// TIA Portal project "PalletizerLine" (V17) (continued)
VERSION : 1.0
// Support: tech.team.motioncontrol@siemens.com
// Fax: +49 (0) 9131/98-1297
   VAR
      Summation : "CPG_typeEventSummation";   // Unit Mode - PackML Event Summation
   END_VAR
BEGIN
   Summation.wrk_EventArraySize := 30;
END_DATA_BLOCK

DATA_BLOCK "PackML"   // DB31613
TITLE = CPG_PackML
{ S7_Optimized_Access := 'TRUE' }
AUTHOR : tech.team.motioncontrol@siemens.com
FAMILY : CPG
VERSION : 1.0
// Support: tech.team.motioncontrol@siemens.com
// Fax: +49 (0) 9131/98-1297
   VAR
      projectVersion : String[10] := 'V1.0.0';   // Project specific version
      Cmd : Struct   // PackML boolean COMMAND to PackML ModeManager & State Model
         Mode : Struct   // Boolean command to change the MODE
            Production : Bool;   // Request to goto mode - PRODUCTION (mode #1)
            Maintenance : Bool;   // Request to goto mode - MAINTENANCE (mode #2)
            Manual : Bool;   // Request to goto mode - MANUAL (mode #3)
            UserMode01 : Bool;   // Request to goto mode - USER MODE 01 (mode #4)
            UserMode02 : Bool;   // Request to goto mode - USER MODE 02 (mode #5)
            UserMode03 : Bool;   // Request to goto mode - USER MODE 03 (mode #6)
            UserMode04 : Bool;   // Request to goto mode - USER MODE 04 (mode #7)
            UserMode05 : Bool;   // Request to goto mode - USER MODE 05 (mode #8)
            UserMode06 : Bool;   // Request to goto mode - USER MODE 06 (mode #9)
            UserMode07 : Bool;   // Request to goto mode - USER MODE 07 (mode #10)
            UserMode08 : Bool;   // Request to goto mode - USER MODE 08 (mode #11)
         END_STRUCT;
      END_STRUCT;
      Sts : Struct   // Status for current mode and state as boolean
         Mode : Struct   // Status of the current MODE
            Production : Bool;   // Current mode - PRODUCTION (mode #1)
            Maintenance : Bool;   // Current mode - MAINTENANCE (mode #2)
            Manual : Bool;   // Current mode - MANUAL (mode #3)
            UserMode01 : Bool;   // Current mode - USER MODE 01 (mode #4)
            UserMode02 : Bool;   // Current mode - USER MODE 02 (mode #5)
            UserMode03 : Bool;   // Current mode - USER MODE 03 (mode #6)
            UserMode04 : Bool;   // Current mode - USER MODE 04 (mode #7)
            UserMode05 : Bool;   // Current mode - USER MODE 05 (mode #8)
            UserMode06 : Bool;   // Current mode - USER MODE 06 (mode #9)
            UserMode07 : Bool;   // Current mode - USER MODE 07 (mode #10)
            UserMode08 : Bool;   // Current mode - USER MODE 08 (mode #11)
         END_STRUCT;
         State : Struct   // Status of the current STATE
            Clearing : Bool;   // Current state is - Clearing
            Stopped : Bool;   // Current state is - Stopped
            Starting : Bool;   // Current state is - Starting
            Idle : Bool;   // Current state is - Idle
            Suspended : Bool;   // Current state is - Suspended
            Execute : Bool;   // Current state is - Executing
            Stopping : Bool;   // Current state is - Stopping
            Aborting : Bool;   // Current state is - Aborting
            Aborted : Bool;   // Current state is - Aborted
            Holding : Bool;   // Current state is - Holding
            Held : Bool;   // Current state is - Held
            Unholding : Bool;   // Current state is - Unholding
            Suspending : Bool;   // Current state is - Suspending
            Unsuspending : Bool;   // Current state is - Unsuspending
            Resetting : Bool;   // Current state is - Resetting
            Completing : Bool;   // Current state is - Completing
            Complete : Bool;   // Current state is - Complete
         END_STRUCT;
      END_STRUCT;
      Cmd_Reset : Bool;   // Request for command - RESET
      Cmd_Start : Bool;   // Request for command - START
      Cmd_Stop : Bool;   // Request for command - STOP
      Cmd_Hold : Bool;   // Request for command - HOLD
      Cmd_UnHold : Bool;   // Request for command - UNHOLD
      Cmd_Suspend : Bool;   // Request for command - SUSPEND
      Cmd_UnSuspend : Bool;   // Request for command - UNSUSPEND
      Cmd_Abort : Bool;   // Request for command - ABORT
      Cmd_Clear : Bool;   // Request for command - CLEAR
      Cmd_Complete : Bool;   // Request for command - COMPLETE
      remoteCommandEnable : Bool;   // If 0 = local mode for PackML commands, if 1=remote command for PackML
      OEE : Struct   // Real-Time OEE values
         realTime : Real;   // Real-Time value (0-100%)
         availability : Real;   // Availability value (0-100%)
         performance : Real;   // Performance value (0-100%)
         quality : Real;   // Quality value (0-100%)
      END_STRUCT;
      PackMLDiag : "typeLPMLV30_Diagnostics";   // PackML Diagnostic Data
   END_VAR
BEGIN
END_DATA_BLOCK

DATA_BLOCK "PackTags"   // DB31614
TITLE = CPG_PackTags
{ S7_Optimized_Access := 'TRUE' }
AUTHOR : tech.team.motioncontrol@siemens.com
FAMILY : CPG
VERSION : 1.0
// Support: tech.team.motioncontrol@siemens.com
// Fax: +49 (0) 9131/98-1297
   VAR
      Command : Struct   // PackTags "Command" tag area. Data is scalable for needs.
         UnitMode : DInt;   // Unit Mode Target (1=Production,2=Maintenance,3=Manual,4=UserMode1,...,31=UserMode28)
         UnitModeChangeRequest : Bool;   // 1=Request Unit Mode Change to commanded value (UnitMode)
         MachSpeed : Real := 0.0;   // Setpoint of Machine Speed in Primary Packages per Minute
         MaterialInterlock : DWord;   // Materials Interlock Command (1=Ready or Not low, 0=Not ready or Low)
         CntrlCmd : DInt;   // State Control Command to drive a state change (1=Reset,2=Start,3=Stop,4=Hold,5=Unhold,6=Suspend,7=Unsuspend,8=Abort,9=Clear)
         CmdChangeRequest : Bool;   // 1=Request Machine State Change to commanded value (CntrlCmd)
         Parameter : Array[0.."CPG_NO_OF_COMMAND_PARAMETERS_UPPER_LIM"] of "CPG_typeParameter(Real)";   // Parameter Structure Array from SCADA / MES
      END_STRUCT;
      Status : Struct   // PackTags "Status" tag area. Data is scalable for needs.
         UnitModeCurrent : DInt := 3;   // Current Unit Mode (1=Production,2=Maintenance,3=Manual,4=UserMode1,...,31=UserMode28)
         UnitModeCurrentName : String[18] := 'Manual';   // Current Unit Mode Name (NOT ISA-TR88 - OPTIONAL)
         UnitModeRequested : Bool;   // 1=Ack. that a unit mode change has been requested
         UnitModeChangeInProcess : Bool;   // 1=Requested Unit Mode Change In Progress
         StateCurrent : DInt := 2;   // Current Machine State (1=Clearing,2=Stopped,3=Starting,4=Idle,5=Suspended,6=Execute,7=Stopping,8=Aborting,9=Aborted,10=Holding,11=Held,12=Unholding,13=Suspending,14=Unsuspending,15=Resetting,16=Completing,17=Complete)
         StateCurrentName : String[16] := 'Stopped';   // Current Machine State name (NOT ISA-TR88 - OPTIONAL)
         StateRequested : DInt;   // Target Machine State
         StateChangeInProcess : Bool;   // 1=Requested State Change in Progress
         MachSpeed : Real := 0.0;   // Setpoint of Machine Speed in Primary Packages per Minute
         CurMachSpeed : Real := 0.0;   // Actual Value of Machine Speed in Primary Packages per Minute
         MaterialInterlock : DWord;   // Materials Interlock Status (1=Ready or Not low, 0=Not ready or Low)
         EquipmentInterlock : Struct   // Machine upstream and downstream status
            Blocked : Bool;   // 1=The downstream system is not able to accept products, 0=all OK
            Starved : Bool;   // 1=The upstream system is not able to supply products, 0=all OK
         END_STRUCT;
         Parameter : Array[0.."CPG_NO_OF_STATUS_PARAMETERS_UPPER_LIM"] of "CPG_typeParameter(Real)";   // Parameter Structure Array for HMI / SCADA / MES
      END_STRUCT;
   END_VAR
   VAR RETAIN
      Admin : Struct   // PackTags "Administration" tag area. Data is scalable for needs.
         Parameter : Array[0.."CPG_NO_OF_ADMIN_PARAMETERS_UPPER_LIM"] of "CPG_typeParameter(Real)";   // Parameter Structure Array for HMI / SCADA / MES
         Alarm : Array[0.."CPG_NO_OF_ADMIN_EVENTS_UPPER_LIM"] of "CPG_typeEvent";   // Alarm summary of Active Events
         AlarmExtent : DInt;   // Number of active alarms
         AlarmHistory : Array[0.."CPG_NO_OF_ADMIN_EVENTS_HISTORY_UPPER_LIM"] of "CPG_typeEvent";   // Alarm History
         AlarmHistoryExtent : DInt;   // Number of alarms in alarm history
         StopReason : "CPG_typeEvent";   // First Fault Alarm Code
         Warning : Array[0.."CPG_NO_OF_ADMIN_EVENTS_UPPER_LIM"] of "CPG_typeEvent";   // Active Machine Warnings
         WarningExtent : DInt;   // Number of Active Machine Warnings
         ModeCurrentTime : Array[0.."LPMLV30_MODES_UPPER_LIM"] of DInt;   // Time spent in the last mode [seconds] (reset each time new mode is entered)
         ModeCumulativeTime : Array[0.."LPMLV30_MODES_UPPER_LIM"] of DInt;   // Cumulative Time for all Modes [seconds]
         StateCurrentTime : Array[0.."LPMLV30_MODES_UPPER_LIM", 0.."LPMLV30_STATES_UPPER_LIM"] of DInt;   // Time spent in the last state [seconds] (reset each time new state is entered)
         StateCumulativeTime : Array[0.."LPMLV30_MODES_UPPER_LIM", 0.."LPMLV30_STATES_UPPER_LIM"] of DInt;   // Cumulative Time for all States [seconds]
         ProdConsumedCount : Array[0.."CPG_NO_OF_PROD_CONSUMED_COUNT_UPPER_LIM"] of "CPG_typeProdCount(DINT)";   // Total Number of Products consumed- good or bad
         ProdProcessedCount : Array[0.."CPG_NO_OF_PROD_PROCESSED_COUNT_UPPER_LIM"] of "CPG_typeProdCount(DINT)";   // Total Number of Products processed - good or bad
         ProdDefectiveCount : Array[0.."CPG_NO_OF_PROD_DEFECTIVE_COUNT_UPPER_LIM"] of "CPG_typeProdCount(DINT)";   // Total Number of Defective (bad) Products processed
         AccTimeSinceLastReset : DInt := L#0;   // Accumulated Time Since Last Reset of all mode and state times and counts
         MachDesignSpeed : Real := 0.0;   // Machine Design Speed of the Current Product Configuration
         StatesDisabled : DInt;   // States 1 to 17 of the PackML State Model can be disabled by turning on the corresponding bit in the DINT
         PLCDateTime : Array[0..6] of DInt;   // Current Date and Time of PLC
         PLCDateTimeDTL : DTL;   // Current Date and LTime (DTL) of PLC (date and time-of-day information in nanoseconds since 01/01/1970 0:0)
      END_STRUCT;
   END_VAR
BEGIN
   Admin.ProdProcessedCount[0]."Name" := 'Processed #1';
   Admin.ProdProcessedCount[0].Unit := 'count';
   Admin.ProdConsumedCount[0]."Name" := 'Consumed #1';
   Admin.ProdConsumedCount[0].Unit := 'count';
   Admin.ProdDefectiveCount[0].Unit := 'count';
   Admin.ProdDefectiveCount[0]."Name" := 'Defective #1';
END_DATA_BLOCK

DATA_BLOCK "HMI_Data"   // DB31615
TITLE = CPG_HMI_Data
{ S7_Optimized_Access := 'TRUE' }
AUTHOR : tech.team.motioncontrol@siemens.com
FAMILY : CPG
VERSION : 1.0
// Support: tech.team.motioncontrol@siemens.com
// Fax: +49 (0) 9131/98-1297
   VAR
      resetPackMLTimers : Bool;   // Reset the PackML Timer values when set (1).
   END_VAR
   VAR RETAIN
      languageSelected : Int;   // This is the value of the language selected in the HMI (0=English, 1=DE, 2=SP, 3
   END_VAR
   VAR
      modeCurrentTime : DInt;   // Time spent in the current mode [seconds](reset each time new mode is entered)
      modeCumulativeTime : DInt;   // Accumulative Time spent in the current mode [seconds]
      State_Current_Times : Array[0.."LPMLV30_STATES_UPPER_LIM"] of DInt;   // Current Time (# of seconds) spent for each state for active mode.
      State_Cumulative_Times : Array[0.."LPMLV30_STATES_UPPER_LIM"] of DInt;   // Accumulative Time (# of seconds) spent for each state for active mode.
      alarmSortedList : Array[0.."CPG_NO_OF_HMI_SORT_EVENTS_UPPER_LIM"] of "CPG_typeEvent";   // Alarm Sorted List for HMI - summary of Active Events
      EM_SortDisable_Alarm : Struct   // Alarm Disable for Equipment Modules (EMs)
         Unit : Bool;   // If bool is reset, then Unit sort filter is enabled, else it's disabled.
         EM00 : Bool;   // If bool is reset, then EMxx sort filter is enabled, else it's disabled.
         EM01 : Bool;   // If bool is reset, then EMxx sort filter is enabled, else it's disabled.
         EM02 : Bool;   // If bool is reset, then EMxx sort filter is enabled, else it's disabled.
         EM03 : Bool;   // If bool is reset, then EMxx sort filter is enabled, else it's disabled.
         EM04 : Bool;   // If bool is reset, then EMxx sort filter is enabled, else it's disabled.
         EM05 : Bool;   // If bool is reset, then EMxx sort filter is enabled, else it's disabled.
         EM06 : Bool;   // If bool is reset, then EMxx sort filter is enabled, else it's disabled.
         EM07 : Bool;   // If bool is reset, then EMxx sort filter is enabled, else it's disabled.
         EM08 : Bool;   // If bool is reset, then EMxx sort filter is enabled, else it's disabled.
         EM09 : Bool;   // If bool is reset, then EMxx sort filter is enabled, else it's disabled.
         EM10 : Bool;   // If bool is reset, then EMxx sort filter is enabled, else it's disabled.
      END_STRUCT;
      alarmFilter : "CPG_typeSortFilter";   // HMI Commands to control the Alarm Sort Filter
      warningSortedList : Array[0.."CPG_NO_OF_HMI_SORT_EVENTS_UPPER_LIM"] of "CPG_typeEvent";   // Warning Sorted List for HMI - summary of Active Events
      EMSortDisableWarning : Struct   // Warning Disable for Equipment Modules (EMs)
         Unit : Bool;   // If bool is reset, then Unit sort filter is enabled, else it's disabled.
         EM00 : Bool;   // If bool is reset, then EMxx sort filter is enabled, else it's disabled.
         EM01 : Bool;   // If bool is reset, then EMxx sort filter is enabled, else it's disabled.
         EM02 : Bool;   // If bool is reset, then EMxx sort filter is enabled, else it's disabled.
         EM03 : Bool;   // If bool is reset, then EMxx sort filter is enabled, else it's disabled.
         EM04 : Bool;   // If bool is reset, then EMxx sort filter is enabled, else it's disabled.
         EM05 : Bool;   // If bool is reset, then EMxx sort filter is enabled, else it's disabled.
         EM06 : Bool;   // If bool is reset, then EMxx sort filter is enabled, else it's disabled.
         EM07 : Bool;   // If bool is reset, then EMxx sort filter is enabled, else it's disabled.
         EM08 : Bool;   // If bool is reset, then EMxx sort filter is enabled, else it's disabled.
         EM09 : Bool;   // If bool is reset, then EMxx sort filter is enabled, else it's disabled.
         EM10 : Bool;   // If bool is reset, then EMxx sort filter is enabled, else it's disabled.
      END_STRUCT;
      WarningFilter : "CPG_typeSortFilter";   // HMI Commands to control the Warning Sort Filter
      HMIWarningMsgScroll : String[40];   // Warning Message - scroll of all active warnings
      ModeNames : Array[0.."LPMLV30_MODES_UPPER_LIM"] of String[18];   // Mode Names for selected language
      StateNames : Array[0.."LPMLV30_STATES_UPPER_LIM"] of String[16];   // State Names for selectecd modes
      PLCDateTime : Struct   // Date Time for WinCC Flexible HMI format
         DATE_TIME : Date_And_Time := DT#12-7-12-18:16:34.356;   // Current Time and Date of PLC
         reserve : Array[0..3] of Byte;   // Filler bytes used to sync HMI clock with PLC clock. Do not change.
      END_STRUCT;
      diagnosticsBufferIndexForHMI : Int;   // Diagnostics to HMI
      diagnosticsBufferEntryForHMI : "typeLPMLV30_DiagnosticsEntry";   // Diagnostics to HMI
      HMICoordination : Word;   // HMI Coordination area pointer: Bit0 = Startup; 1=OpMode (0=on, 1=off-line), 2=life bit
      HMICurrentScreenID : Int;   // HMI Current screen number
      CMDs : Struct   // HMI Commands
         PB_Start : Bool;   // HMI Push Button Command - Start
         PB_Stop : Bool;   // HMI Push Button Command - Stop
         PB_Hold : Bool;   // HMI Push Button Command - Hold
         PB_Reset : Bool;   // HMI Push Button Command - Reset
         PB_Complete : Bool;   // HMI Push Button Command - Complete (demo purposes only)
         PB_EStop : Bool;   // HMI Push Button Command - EStop (demo purposes only)
         PB_Abort : Bool;   // HMI Push Button Command - Abort (demo purposes only)
         PB_ProdSimulate : Bool;   // HMI Push Button Command - Product Simulate Enable (demo purposes only)
         PB_DriveSimulate : Bool;   // HMI Push Button Command - Drive / Axis Simulate (demo purposes only)
      END_STRUCT;
   END_VAR
BEGIN
END_DATA_BLOCK

DATA_BLOCK "HMI_Data_Custom"   // DB31616
TITLE = CPG_HMI_Data_Custom
{ S7_Optimized_Access := 'TRUE' }
AUTHOR : tech.team.motioncontrol@siemens.com
FAMILY : CPG
VERSION : 1.0
// Support: tech.team.motioncontrol@siemens.com
// Fax: +49 (0) 9131/98-1297
   VAR
      machineSpeedSP : Real := 20.0;   // Machine Speed Setpoint (product per min)
      machineSpeedPV : Real;   // Machine Speed Actual (product per min)
   END_VAR
BEGIN
END_DATA_BLOCK

DATA_BLOCK "ParetoData"   // DB31617
TITLE = CPG_ParetoData
{ S7_Optimized_Access := 'TRUE' }
AUTHOR : tech.team.motioncontrol@siemens.com
FAMILY : CPG
VERSION : 1.1
// Support: tech.team.motioncontrol@siemens.com
   VAR RETAIN
      alarmOccurrence : Array[0.."CPG_PARTEO_NO_OF_ERRORS_UPPER_LIM"] of "CPG_typePareto";   // Alarm Array
      totalStops : Int;   // Total stops on the machine
      totalTimeSinceReset : Real;   // Total time since reset
      totalUptime : Real;   // Total uptime of the machine
      totalDowntime : Real;   // Total downtime of the machine
      percentUptime : Real;
      MTTR : Real;
      MTBF : Real;
      Sort : Int;
      Reset : Bool;
   END_VAR
BEGIN
END_DATA_BLOCK

DATA_BLOCK "RecipeManagement"   // DB31618
TITLE = CPG_RecipeManagement
{ S7_Optimized_Access := 'TRUE' }
AUTHOR : tech.team.motioncontrol@siemens.com
FAMILY : CPG
VERSION : 1.1
// Support: tech.team.motioncontrol@siemens.com
   VAR
      HMI_Command : Struct   // Helper bits for HMI Recipe Control
         Change : Struct
            changeCmd : Bool;
            changeID : Int;
            cancel : Bool;
            request : Bool;
         END_STRUCT;
         Save : Struct
            saveCmd : Bool;
            saveAsCmd : Bool;
            saveAsDestinationID : Int;
            saveAsNewName : String[60];
            cancel : Bool;
            request : Bool;
         END_STRUCT;
         Copy : Struct
            copyCmd : Bool;
            copySourceID : Int;
            copyDestinationID : Int;
            copyNewName : String[60];
            cancel : Bool;
            request : Bool;
         END_STRUCT;
         Delete : Struct
            deleteCmd : Bool;
            deleteID : Int;
            cancel : Bool;
            request : Bool;
         END_STRUCT;
         resetAllTimes : Bool;
      END_STRUCT;
      HMI_Indicator : Struct   // Helper bits for HMI Recipe Control
         changeConfirm : Bool;
         saveAsConfirm : Bool;
         copyConfirm : Bool;
         deleteConfirm : Bool;
         changeErr : Bool;
         saveAsErr : Bool;
         copyErr : Bool;
         deleteErr : Bool;
      END_STRUCT;
      setpointsArray_REAL : Array[0..11] of "CPG_typeRecipeSetpoint_REAL";   // The setpoints that are displayed
      setpointsArray_DINT : Array[0..11] of "CPG_typeRecipeSetpoint_DINT";   // The setpoints that are displayed
      setpointsArray_BOOL : Array[0..11] of "CPG_typeRecipeSetpoint_BOOL";   // The setpoints that are displayed
      setpointsArray_STRING : Array[0..11] of "CPG_typeRecipeSetpoint_STRING";   // The setpoints that are displayed
      setpointPopup_REAL : "CPG_typeRecipeSetpoint_REAL";   // The setpoint in the popup
      setpointPopup_DINT : "CPG_typeRecipeSetpoint_DINT";   // The setpoint in the popup
      setpointPopup_BOOL : "CPG_typeRecipeSetpoint_BOOL";   // The setpoint in the popup
      setpointPopup_STRING : "CPG_typeRecipeSetpoint_STRING";   // The setpoint in the popup
      popupTrackers : Array[0..3] of Int;   // Int to track the location of popup
      currentPages : Array[0..4] of Int;   // Current page of setpoints (or recipes)
      maxPages : Array[0..4] of Int;   // Max page of setpoints (or recipes)
      displayDisable_REAL : Array[0..11] of Bool;   // True if that setpoint should be hidden
      displayDisable_DINT : Array[0..11] of Bool;   // True if that setpoint should be hidden
      displayDisable_BOOL : Array[0..11] of Bool;   // True if that setpoint should be hidden
      displayDisable_STRING : Array[0..11] of Bool;   // True if that setpoint should be hidden
      recipeArrayNames : Array[0..19] of String[60];   // Recipe names to display
      recipeArraySaves : Array[0..19] of DTL;   // Recipe times to display
      recipeArrayTimes : Array[0..19] of Time;   // Recipe savepoints to display
      recipeArrayNums : Array[0..19] of Int;   // Recipe numbers
      recipeArrayHide : Array[0..19] of Bool;   // True if that recipe should be hidden
   END_VAR
BEGIN
   currentPages[0] := 1;
   currentPages[2] := 1;
   currentPages[1] := 1;
   currentPages[3] := 1;
   maxPages[0] := 1;
   maxPages[2] := 1;
   maxPages[3] := 1;
   maxPages[1] := 1;
   currentPages[4] := 1;
END_DATA_BLOCK

// folder: GlobalData/Configuration

DATA_BLOCK "RecipeCfg"   // DB1605
TITLE = CPG_RecipeCfg
{ S7_Optimized_Access := 'TRUE' }
AUTHOR : tech.team.motioncontrol@siemens.com
FAMILY : CPG
VERSION : 1.1
// Support: tech.team.motioncontrol@siemens.com
   VAR
      setpoints_REAL : Array[0.."CPG_NO_OF_SETPOINT_REAL_UPPER_LIM"] of "CPG_typeRecipeSetpoint_REAL";   // Array of setpoints of REAL
      setpoints_DINT : Array[0.."CPG_NO_OF_SETPOINT_DINT_UPPER_LIM"] of "CPG_typeRecipeSetpoint_DINT";   // Array of setpoints of DINT
      setpoints_BOOL : Array[0.."CPG_NO_OF_SETPOINT_BOOL_UPPER_LIM"] of "CPG_typeRecipeSetpoint_BOOL";   // Array of setpoints of BOOL
      setpoints_STRING : Array[0.."CPG_NO_OF_SETPOINT_STRING_UPPER_LIM"] of "CPG_typeRecipeSetpoint_STRING";   // Array of setpoints of STRING
      recipeControl : "CPG_typeRecipeControl";   // FB_Recipe_Control communicates to the setpoints via this tag
      recipeNames : Array[0.."CPG_NO_OF_RECIPE_UPPER_LIM"] of String[60];   // Array holding the names of all recipes
      recipeCumTimes : Array[0.."CPG_NO_OF_RECIPE_UPPER_LIM"] of Time;   // Array holding the cumulative time all recipes have been active
      recipeLastSaveTimes : Array[0.."CPG_NO_OF_RECIPE_UPPER_LIM"] of DTL;   // Array holding the last time each recipe was saved
   END_VAR
BEGIN
   recipeNames[0] := 'Recipe 0';
   recipeNames[1] := 'Recipe 1';
   recipeNames[2] := 'Recipe 2';
   recipeNames[3] := 'Recipe 3';
   recipeNames[4] := 'Recipe 4';
   recipeNames[5] := 'Recipe 5';
   recipeNames[6] := 'Recipe 6';
   recipeNames[7] := 'Recipe 7';
   recipeNames[8] := 'Recipe 8';
   recipeNames[9] := 'Recipe 9';
   recipeNames[10] := 'Recipe 10';
   recipeNames[11] := 'Recipe 11';
   recipeNames[12] := 'Recipe 12';
   recipeNames[13] := 'Recipe 13';
   recipeControl.RecipeID_A := 1;
   recipeControl.RecipeID_B := 2;
   recipeControl.RecipeID_C := 3;
   setpoints_BOOL[0].Text_True[0] := 'TRUE';
   setpoints_BOOL[0].SetpointName[1] := '';
   setpoints_BOOL[0].SetpointName[0] := 'BOOL SP 0';
   recipeNames[14] := 'Recipe 14';
   recipeNames[15] := 'Recipe 15';
   recipeNames[16] := 'Recipe 16';
   recipeNames[17] := 'Recipe 17';
   recipeNames[18] := 'Recipe 18';
   recipeNames[19] := 'Recipe 19';
   recipeNames[20] := 'Recipe 20';
   recipeControl.CurrentRecipeID := 0;
   recipeControl.CurrentRecipeName := 'Recipe 0';
   recipeLastSaveTimes[0] := DTL#2019-1-1-00:00:00;
   recipeLastSaveTimes[1] := DTL#2019-1-1-00:00:00;
   recipeLastSaveTimes[2] := DTL#2019-1-1-00:00:00;
   recipeLastSaveTimes[3] := DTL#2019-1-1-00:00:00;
   recipeLastSaveTimes[4] := DTL#2019-1-1-00:00:00;
   recipeLastSaveTimes[5] := DTL#2019-1-1-00:00:00;
   recipeLastSaveTimes[6] := DTL#2019-1-1-00:00:00;
   recipeLastSaveTimes[7] := DTL#2019-1-1-00:00:00;
   recipeLastSaveTimes[8] := DTL#2019-1-1-00:00:00;
   recipeLastSaveTimes[9] := DTL#2019-1-1-00:00:00;
   recipeLastSaveTimes[10] := DTL#2019-1-1-00:00:00;
   recipeLastSaveTimes[11] := DTL#2019-1-1-00:00:00;
   recipeLastSaveTimes[12] := DTL#2019-1-1-00:00:00;
   recipeLastSaveTimes[13] := DTL#2019-1-1-00:00:00;
   recipeLastSaveTimes[14] := DTL#2019-1-1-00:00:00;
   recipeLastSaveTimes[15] := DTL#2019-1-1-00:00:00;
   recipeLastSaveTimes[16] := DTL#2019-1-1-00:00:00;
   recipeLastSaveTimes[17] := DTL#2019-1-1-00:00:00;
   recipeLastSaveTimes[18] := DTL#2019-1-1-00:00:00;
   recipeLastSaveTimes[19] := DTL#2019-1-1-00:00:00;
   recipeLastSaveTimes[20] := DTL#2019-1-1-00:00:00;
   setpoints_DINT[0].SetpointName[0] := 'DINT SP 0';
   setpoints_REAL[0].SetpointName[0] := 'LH 1 Length';
   setpoints_BOOL[0].Text_True[1] := '';
   setpoints_BOOL[0].Text_False[0] := 'FALSE';
   setpoints_STRING[0].SetpointName[0] := 'STRING SP 0';
   setpoints_STRING[0].RecipeValues[0] := 'a';
   setpoints_STRING[0].RecipeValues[1] := 'b';
   setpoints_STRING[0].RecipeValues[2] := 'c';
   setpoints_STRING[0].RecipeValues[3] := 'd';
   setpoints_STRING[0].RecipeValues[4] := 'e';
   setpoints_STRING[0].RecipeValues[5] := 'f';
   setpoints_STRING[0].RecipeValues[6] := 'g';
END_DATA_BLOCK

DATA_BLOCK "AlarmCfg"   // DB31600
TITLE = CPG_AlarmCfg
{ S7_Optimized_Access := 'TRUE' }
AUTHOR : tech.team.motioncontrol@siemens.com
FAMILY : CPG
VERSION : 1.0
// Support: tech.team.motioncontrol@siemens.com
// Fax: +49 (0) 9131/98-1297
   VAR
      Event : Array[0.."CPG_NO_OF_CFG_ALARMS_UPPER_LIM"] of "CPG_typeEventCfg";
   END_VAR
BEGIN
   Event[0].ID := 0;
   Event[0].category := 6;
   Event[0].message[0] := 'Alarm Test';
   Event[0].message[1] := 'Alarm Test';
   Event[1].message[0] := 'E-Stop';
   Event[1].message[1] := 'Not-Halt';
   Event[1].ID := 1;
   Event[1].value := 1;
   Event[1].category := 0;   // 0 = Safety related, Coordinated fast stop
   Event[2].message[0] := 'Guard Door';
   Event[2].message[1] := 'Schutzzaun';
   Event[2].ID := 4;
   Event[2].value := 1;
   Event[3].ID := 33;
   Event[3].value := 2;
   Event[3].message[0] := 'Stop PB';
   Event[3].message[1] := 'Stopp Taster';
   Event[3].category := 2;   // 2 = Coordinated normal stop
   Event[4].message[0] := 'Hold PB';
   Event[4].message[1] := 'Hold Taster';
   Event[4].ID := 40;
   Event[4].value := 0;
   Event[4].category := 7;   // 7 = Held command
   Event[5].ID := 262;
   Event[5].value := 0;
   Event[5].category := 1;   // 1 = Coordinated fast stop
   Event[5].message[0] := 'Axis Error';
   Event[5].message[1] := 'Achsfehler';
   Event[6].ID := 261;
   Event[6].value := 1;
   Event[6].category := 1;   // 1 = Coordinated fast stop
   Event[6].message[0] := 'Drive Faulted';
   Event[6].message[1] := 'Antriebsfehler';
   Event[7].ID := 7;
   Event[7].value := 7;
   Event[7].category := 8;   // 8 =Blocked, Coordinated slow stop
   Event[7].message[0] := 'Machine Blocked';
   Event[7].message[1] := 'Maschine blockiert';
   Event[8].message[0] := 'Starved - No botttles';
   Event[8].message[1] := 'Flaschenzufuhr leer';
   Event[8].category := 9;   // 9 = Starved, Coordinated slow stop
   Event[8].ID := 8;
   Event[8].value := 8;
   Event[9].message[0] := 'Starved - No labels';
   Event[9].message[1] := 'Etikettenzufuhr leer';
   Event[9].category := 9;   // 9 = Starved, Coordinated slow stop
   Event[9].ID := 9;
   Event[9].value := 9;
   Event[10].message[0] := 'Spare';
   Event[10].message[1] := 'Reserve';
   Event[10].category := 0;   // 9 = Starved, Coordinated slow stop
   Event[11].message[0] := 'Spare';
   Event[11].message[1] := 'Reserve';
   Event[11].category := 0;
   Event[12].message[0] := 'Spare';
   Event[12].message[1] := 'Reserve';
   Event[12].category := 0;
   Event[13].message[0] := 'Spare';
   Event[13].message[1] := 'Reserve';
   Event[13].category := 0;
   Event[14].message[0] := 'Spare';
   Event[14].message[1] := 'Reserve';
   Event[15].message[0] := 'Spare';
   Event[15].message[1] := 'Reserve';
   Event[16].message[0] := 'Spare';
   Event[16].message[1] := 'Reserve';
   Event[17].message[0] := 'Spare';
   Event[17].message[1] := 'Reserve';
   Event[18].message[0] := 'Spare';
   Event[18].message[1] := 'Reserve';
   Event[19].message[0] := 'Spare';
   Event[19].message[1] := 'Reserve';
   Event[20].message[0] := 'Remote Stop Cmd';
   Event[20].message[1] := 'Remote Stop Cmd';
   Event[20].ID := 41;
   Event[20].value := 20;
   Event[20].category := 2;   // 2 = Coordinated normal stop
   Event[21].message[0] := 'Remote Abort Cmd';
   Event[21].message[1] := 'Remote Abort Cmd';
   Event[21].ID := 42;
   Event[21].value := 21;
   Event[22].ID := 43;
   Event[22].value := 22;
   Event[22].message[0] := 'Rmt Suspd Cmd - Blocked';
   Event[22].message[1] := 'Remote Suspend Cmd - Blocked';
   Event[22].category := 8;   // 9 = Starved, Coordinated slow stop
   Event[23].message[0] := 'Rmt Suspd Cmd - Starved';
   Event[23].message[1] := 'Remote Suspend Cmd - Starved';
   Event[23].category := 9;   // 7 = Hold, Coordinated slow stop
   Event[23].ID := 43;
   Event[23].value := 23;
   Event[24].message[0] := 'Remote Hold Cmd';
   Event[24].message[1] := 'Remote Hold Cmd';
   Event[21].category := 1;   // 0 = Safety related, Coordinated fast stop
   Event[25].message[0] := 'Spare';
   Event[25].message[1] := 'Reserve';
   Event[26].message[0] := 'Spare';
   Event[26].message[1] := 'Reserve';
   Event[27].message[0] := 'Spare';
   Event[27].message[1] := 'Reserve';
   Event[28].message[0] := 'Spare';
   Event[28].message[1] := 'Reserve';
   Event[29].message[0] := 'Spare';
   Event[29].message[1] := 'Reserve';
   Event[30].message[0] := 'Spare';
   Event[30].message[1] := 'Reserve';
   Event[31].message[1] := 'Reserve';
   Event[31].message[0] := 'Spare';
   Event[24].ID := 44;
   Event[24].value := 24;
   Event[24].category := 7;   // 7 = Coordinated slow stop
   Event[39].message[1] := 'Reserve';
   Event[39].message[0] := 'Spare';
   Event[38].message[1] := 'Reserve';
   Event[38].message[0] := 'Spare';
   Event[38].value := 0;
   Event[37].message[1] := 'Reserve';
   Event[37].message[0] := 'Spare';
   Event[36].message[1] := 'Reserve';
   Event[36].message[0] := 'Spare';
   Event[35].message[1] := 'Reserve';
   Event[35].message[0] := 'Spare';
   Event[34].message[1] := 'Reserve';
   Event[34].message[0] := 'Spare';
   Event[33].message[1] := 'Reserve';
   Event[33].message[0] := 'Spare';
   Event[32].message[1] := 'Reserve';
   Event[32].message[0] := 'Spare';
   Event[0].message[2] := 'Alarm Test';
   Event[1].message[2] := 'Los E-Stop';
   Event[2].message[2] := 'Las Guard Door';
   Event[3].message[2] := 'Las Stop PB';
   Event[4].message[2] := 'Las Hold PB';
   Event[5].message[2] := 'Las Axis Error';
   Event[6].message[2] := 'Los Drive Faulted';
   Event[7].message[2] := 'Los Machine Blocked';
   Event[8].message[2] := 'Las Starved - No botttles';
   Event[9].message[2] := 'Las Starved - No labels';
   Event[10].message[2] := 'Spare';
   Event[11].message[2] := 'Spare';
   Event[12].message[2] := 'Spare';
   Event[13].message[2] := 'Spare';
   Event[14].message[2] := 'Spare';
   Event[15].message[2] := 'Spare';
   Event[16].message[2] := 'Spare';
   Event[17].message[2] := 'Spare';
   Event[18].message[2] := 'Spare';
   Event[19].message[2] := 'Spare';
   Event[20].message[2] := 'Las Remote Stop Cmd';
   Event[21].message[2] := 'Las Remote Abort Cmd';
   Event[22].message[2] := 'Las Remote Suspd Cmd - Blocked';
   Event[23].message[2] := 'Las Rmt Suspd Cmd - Starved';
   Event[24].message[2] := 'Las Remote Hold Cmd';
   Event[25].message[2] := 'Spare';
   Event[26].message[2] := 'Spare';
   Event[27].message[2] := 'Spare';
   Event[28].message[2] := 'Spare';
   Event[29].message[2] := 'Spare';
   Event[30].message[2] := 'Spare';
   Event[31].message[2] := 'Spare';
   Event[32].message[2] := 'Spare';
   Event[33].message[2] := 'Spare';
   Event[34].message[2] := 'Spare';
   Event[35].message[2] := 'Spare';
   Event[36].message[2] := 'Spare';
   Event[37].message[2] := 'Spare';
   Event[38].message[2] := 'Spare';
   Event[39].message[2] := 'Spare';
   // Event[0] : Alarm Test
   // Event[1] : Emergency Stop
   // Event[2] : Guard Door
   // Event[2].category : 0 = Safety related, Coordinated fast stop
   // Event[3] : Stop Command
   // Event[4] : Hold Command
   // Event[5] : Axis Error
   // Event[6] : Drive Fault
   // Event[7] : Machine Blocked
   // Event[8] : Machine Starved - No bottles
   // Event[9] : Machine Starved - No labels
   // Event[10] : Spare
   // Event[11] : Spare
   // Event[12] : Spare
   // Event[13] : Spare
   // Event[14] : Spare
   // Event[15] : Spare
   // Event[16] : Spare
   // Event[17] : Spare
   // Event[18] : Spare
   // Event[19] : Spare
   // Event[20] : Remote Stop Command
   // Event[21] : Remote Abort Command
   // Event[22] : Rmt Suspd Cmd - Blocked
   // Event[23] : Rmt Suspd Cmd - Starved
   // Event[24] : Remote Hold Cmd
   // Event[25] : Spare
   // Event[26] : Spare
   // Event[27] : Spare
   // Event[28] : Spare
   // Event[29] : Spare
   // Event[31] : Spare
   // Event[30] : Spare
   // Event[32] : Spare
   // Event[33] : Spare
   // Event[34] : Spare
   // Event[35] : Spare
   // Event[36] : Spare
   // Event[37] : Spare
   // Event[38] : Spare
   // Event[39] : Spare
END_DATA_BLOCK

DATA_BLOCK "StatusCfg"   // DB31602
TITLE = CPG_StatusCfg
{ S7_Optimized_Access := 'TRUE' }
AUTHOR : tech.team.motioncontrol@siemens.com
FAMILY : CPG
VERSION : 1.0
// Support: tech.team.motioncontrol@siemens.com
// Fax: +49 (0) 9131/98-1297
   VAR
      Event : Array[0.."CPG_NO_OF_CFG_STATUS_UPPER_LIM"] of "CPG_typeEventCfg";
   END_VAR
BEGIN
   Event[0].message[0] := 'Status Test';
   Event[0].message[1] := 'Status Test';
   Event[1].ID := 1;
   Event[1].message[0] := 'Alarms Present';
   Event[2].message[0] := 'Waiting for Reset PB';
   Event[2].message[1] := 'Warte auf Reset Taste';
   Event[1].message[1] := 'Alarme anstehend';
   Event[3].message[0] := 'Waiting for Start PB';
   Event[3].message[1] := 'Warten auf Start Taste';
   Event[4].message[0] := 'Not Ready for Motion';
   Event[4].message[1] := 'Maschine nicht anlaufbereit';
   Event[5].message[0] := 'Waiting for No Motion';
   Event[5].message[1] := 'Warte auf Maschinenstillstand';
   Event[6].message[0] := 'Waiting to start Gearing';
   Event[7].message[0] := 'Waiting to Finish';
   Event[7].message[1] := 'Warte auf Ende Leerfahren';
   Event[8].message[0] := 'Waiting for Un-Hold PB';
   Event[8].message[1] := 'Warte auf Un-Hold Taste';
   Event[9].message[0] := 'Waiting for Mat. Supply';
   Event[9].message[1] := 'Warte auf Materialversorgung';
   Event[10].message[0] := 'Spare';
   Event[10].message[1] := 'Reserve';
   Event[11].message[0] := 'Spare';
   Event[11].message[1] := 'Reserve';
   Event[12].message[0] := 'Spare';
   Event[12].message[1] := 'Reserve';
   Event[13].message[1] := 'Reserve';
   Event[13].message[0] := 'Spare';
   Event[14].message[0] := 'Spare';
   Event[14].message[1] := 'Reserve';
   Event[15].message[0] := 'Spare';
   Event[15].message[1] := 'Reserve';
   Event[16].message[0] := 'Spare';
   Event[16].message[1] := 'Reserve';
   Event[18].message[0] := 'Spare';
   Event[18].message[1] := 'Reserve';
   Event[19].message[1] := 'Reserve';
   Event[19].message[0] := 'Spare';
   Event[0].ID := 0;
   Event[2].ID := 2;
   Event[3].ID := 3;
   Event[4].ID := 4;
   Event[5].ID := 5;
   Event[6].ID := 6;
   Event[7].ID := 7;
   Event[8].ID := 8;
   Event[9].ID := 9;
   Event[10].ID := 10;
   Event[11].ID := 11;
   Event[12].ID := 12;
   Event[13].ID := 13;
   Event[14].ID := 14;
   Event[15].ID := 15;
   Event[16].ID := 16;
   Event[17].ID := 17;
   Event[18].ID := 18;
   Event[19].ID := 19;
   Event[0].message[2] := 'Los Status Test';
   Event[1].message[2] := 'Las Alarms Present';
   Event[2].message[2] := 'Esperando de Reajustar PB';
   Event[3].message[2] := 'Esperando de Comenzar PB';
   Event[4].message[2] := 'No Listo para Movimiento';
   Event[5].message[2] := 'Esperando No Movimiento';
   Event[6].message[2] := 'Waiting to start Gearing';
   Event[6].message[1] := 'Warte auf Start Getriebegleichlauf';
   Event[7].message[2] := 'Esperando para Terminar';
   Event[8].message[2] := 'Waiting for Un-Hold PB';
   Event[9].message[2] := 'Waiting for Mat. Supply';
   Event[10].message[2] := 'Spare';
   Event[11].message[2] := 'Spare';
   Event[12].message[2] := 'Spare';
   Event[13].message[2] := 'Spare';
   Event[14].message[2] := 'Spare';
   Event[15].message[2] := 'Spare';
   Event[16].message[2] := 'Spare';
   Event[17].message[0] := 'Spare';
   Event[17].message[1] := 'Reserve';
   Event[17].message[2] := 'Spare';
   Event[18].message[2] := 'Spare';
   Event[19].message[2] := 'Spare';
   // Event[0] : Status Test
   // Event[1] : 'Alarms Present'
   // Event[2] : 'Waiting for Reset Cmd'
   // Event[3] : 'Waiting for Start Cmd'
   // Event[4] : 'Not Ready for Motion'
   // Event[5] : 'Waiting for No Motion'
   // Event[6] : 'Waiting to start Gearing'
   // Event[7] : 'Waiting to Finish'
   // Event[8] : 'Waiting for Un-Hold Cmd'
   // Event[9] : 'Waiting for Mat. Supply'
   // Event[10] : Spare
   // Event[11] : Spare
   // Event[12] : Spare
   // Event[13] : Spare
   // Event[14] : Spare
   // Event[15] : Spare
   // Event[16] : Spare
   // Event[17] : Spare
   // Event[18] : Spare
   // Event[19] : Spare
END_DATA_BLOCK

DATA_BLOCK "PackMLCfg"   // DB31603
TITLE = CPG_PackMLCfg
{ S7_Optimized_Access := 'TRUE' }
AUTHOR : tech.team.motioncontrol@siemens.com
FAMILY : CPG
VERSION : 1.0
// Support: tech.team.motioncontrol@siemens.com
// Fax: +49 (0) 9131/98-1297
   VAR
      Cfg : "typeLPMLV30_Configuration";   // PackML Configuration Data
      Names : "typeLPMLV30_NamesConfiguration";   // PackML Names Data
      disable : Struct   // Bits used to disable TR88 UN & EMs
         UN : Bool;   // UN (1 = disable, 0= enable)
         EM00 : Struct   // EM00 (1 = disable, 0 = enable)
            EM : Bool;   // EMxx (1 = disable, 0 = enable)
            CM01 : Bool;   // CMxx (1 = disable, 0 = enable)
            CM02 : Bool;   // CMxx (1 = disable, 0 = enable)
            CM03 : Bool;   // CMxx (1 = disable, 0 = enable)
            CM04 : Bool;   // CMxx (1 = disable, 0 = enable)
            CM05 : Bool;   // CMxx (1 = disable, 0 = enable)
            CM06 : Bool;   // CMxx (1 = disable, 0 = enable)
            CM07 : Bool;   // CMxx (1 = disable, 0 = enable)
            CM08 : Bool;   // CMxx (1 = disable, 0 = enable)
            CM09 : Bool;   // CMxx (1 = disable, 0 = enable)
            CM10 : Bool;   // CMxx (1 = disable, 0 = enable)
         END_STRUCT;
         EM01 : Struct   // EM01 (1 = disable, 0 = enable)
            EM : Bool;   // EMxx (1 = disable, 0 = enable)
            CM01 : Bool;   // CMxx (1 = disable, 0 = enable)
            CM02 : Bool;   // CMxx (1 = disable, 0 = enable)
            CM03 : Bool;   // CMxx (1 = disable, 0 = enable)
            CM04 : Bool;   // CMxx (1 = disable, 0 = enable)
            CM05 : Bool;   // CMxx (1 = disable, 0 = enable)
            CM06 : Bool;   // CMxx (1 = disable, 0 = enable)
            CM07 : Bool;   // CMxx (1 = disable, 0 = enable)
            CM08 : Bool;   // CMxx (1 = disable, 0 = enable)
            CM09 : Bool;   // CMxx (1 = disable, 0 = enable)
            CM10 : Bool;   // CMxx (1 = disable, 0 = enable)
         END_STRUCT;
         EM02 : Struct   // EM02 (1 = disable, 0 = enable)
            EM : Bool;   // EMxx (1 = disable, 0 = enable)
            CM01 : Bool;   // CMxx (1 = disable, 0 = enable)
            CM02 : Bool;   // CMxx (1 = disable, 0 = enable)
            CM03 : Bool;   // CMxx (1 = disable, 0 = enable)
            CM04 : Bool;   // CMxx (1 = disable, 0 = enable)
            CM05 : Bool;   // CMxx (1 = disable, 0 = enable)
            CM06 : Bool;   // CMxx (1 = disable, 0 = enable)
            CM07 : Bool;   // CMxx (1 = disable, 0 = enable)
            CM08 : Bool;   // CMxx (1 = disable, 0 = enable)
            CM09 : Bool;   // CMxx (1 = disable, 0 = enable)
            CM10 : Bool;   // CMxx (1 = disable, 0 = enable)
         END_STRUCT;
         EM03 : Struct   // EM03 (1 = disable, 0 = enable)
            EM : Bool;   // EMxx (1 = disable, 0 = enable)
            CM01 : Bool;   // CMxx (1 = disable, 0 = enable)
            CM02 : Bool;   // CMxx (1 = disable, 0 = enable)
            CM03 : Bool;   // CMxx (1 = disable, 0 = enable)
            CM04 : Bool;   // CMxx (1 = disable, 0 = enable)
            CM05 : Bool;   // CMxx (1 = disable, 0 = enable)
            CM06 : Bool;   // CMxx (1 = disable, 0 = enable)
            CM07 : Bool;   // CMxx (1 = disable, 0 = enable)
            CM08 : Bool;   // CMxx (1 = disable, 0 = enable)
            CM09 : Bool;   // CMxx (1 = disable, 0 = enable)
            CM10 : Bool;   // CMxx (1 = disable, 0 = enable)
         END_STRUCT;
         EM04 : Struct   // EM04 (1 = disable, 0 = enable)
            EM : Bool;   // EMxx (1 = disable, 0 = enable)
            CM01 : Bool;   // CMxx (1 = disable, 0 = enable)
            CM02 : Bool;   // CMxx (1 = disable, 0 = enable)
            CM03 : Bool;   // CMxx (1 = disable, 0 = enable)
            CM04 : Bool;   // CMxx (1 = disable, 0 = enable)
            CM05 : Bool;   // CMxx (1 = disable, 0 = enable)
            CM06 : Bool;   // CMxx (1 = disable, 0 = enable)
            CM07 : Bool;   // CMxx (1 = disable, 0 = enable)
            CM08 : Bool;   // CMxx (1 = disable, 0 = enable)
            CM09 : Bool;   // CMxx (1 = disable, 0 = enable)
            CM10 : Bool;   // CMxx (1 = disable, 0 = enable)
         END_STRUCT;
         EM05 : Struct   // EM05 (1 = disable, 0 = enable)
            EM : Bool;   // EMxx (1 = disable, 0 = enable)
            CM01 : Bool;   // CMxx (1 = disable, 0 = enable)
            CM02 : Bool;   // CMxx (1 = disable, 0 = enable)
            CM03 : Bool;   // CMxx (1 = disable, 0 = enable)
            CM04 : Bool;   // CMxx (1 = disable, 0 = enable)
            CM05 : Bool;   // CMxx (1 = disable, 0 = enable)
            CM06 : Bool;   // CMxx (1 = disable, 0 = enable)
            CM07 : Bool;   // CMxx (1 = disable, 0 = enable)
            CM08 : Bool;   // CMxx (1 = disable, 0 = enable)
            CM09 : Bool;   // CMxx (1 = disable, 0 = enable)
            CM10 : Bool;   // CMxx (1 = disable, 0 = enable)
         END_STRUCT;
         EM06 : Struct   // EM06 (1 = disable, 0 = enable)
            EM : Bool;   // EMxx (1 = disable, 0 = enable)
            CM01 : Bool;   // CMxx (1 = disable, 0 = enable)
            CM02 : Bool;   // CMxx (1 = disable, 0 = enable)
            CM03 : Bool;   // CMxx (1 = disable, 0 = enable)
            CM04 : Bool;   // CMxx (1 = disable, 0 = enable)
            CM05 : Bool;   // CMxx (1 = disable, 0 = enable)
            CM06 : Bool;   // CMxx (1 = disable, 0 = enable)
            CM07 : Bool;   // CMxx (1 = disable, 0 = enable)
            CM08 : Bool;   // CMxx (1 = disable, 0 = enable)
            CM09 : Bool;   // CMxx (1 = disable, 0 = enable)
            CM10 : Bool;   // CMxx (1 = disable, 0 = enable)
         END_STRUCT;
         EM07 : Struct   // EM07 (1 = disable, 0 = enable)
            EM : Bool;   // EMxx (1 = disable, 0 = enable)
            CM01 : Bool;   // CMxx (1 = disable, 0 = enable)
            CM02 : Bool;   // CMxx (1 = disable, 0 = enable)
            CM03 : Bool;   // CMxx (1 = disable, 0 = enable)
            CM04 : Bool;   // CMxx (1 = disable, 0 = enable)
            CM05 : Bool;   // CMxx (1 = disable, 0 = enable)
            CM06 : Bool;   // CMxx (1 = disable, 0 = enable)
            CM07 : Bool;   // CMxx (1 = disable, 0 = enable)
            CM08 : Bool;   // CMxx (1 = disable, 0 = enable)
            CM09 : Bool;   // CMxx (1 = disable, 0 = enable)
            CM10 : Bool;   // CMxx (1 = disable, 0 = enable)
         END_STRUCT;
         EM08 : Struct   // EM08 (1 = disable, 0 = enable)
            EM : Bool;   // EMxx (1 = disable, 0 = enable)
            CM01 : Bool;   // CMxx (1 = disable, 0 = enable)
            CM02 : Bool;   // CMxx (1 = disable, 0 = enable)
            CM03 : Bool;   // CMxx (1 = disable, 0 = enable)
            CM04 : Bool;   // CMxx (1 = disable, 0 = enable)
            CM05 : Bool;   // CMxx (1 = disable, 0 = enable)
            CM06 : Bool;   // CMxx (1 = disable, 0 = enable)
            CM07 : Bool;   // CMxx (1 = disable, 0 = enable)
            CM08 : Bool;   // CMxx (1 = disable, 0 = enable)
            CM09 : Bool;   // CMxx (1 = disable, 0 = enable)
            CM10 : Bool;   // CMxx (1 = disable, 0 = enable)
         END_STRUCT;
         EM09 : Struct   // EM09 (1 = disable, 0 = enable)
            EM : Bool;   // EMxx (1 = disable, 0 = enable)
            CM01 : Bool;   // CMxx (1 = disable, 0 = enable)
            CM02 : Bool;   // CMxx (1 = disable, 0 = enable)
            CM03 : Bool;   // CMxx (1 = disable, 0 = enable)
            CM04 : Bool;   // CMxx (1 = disable, 0 = enable)
            CM05 : Bool;   // CMxx (1 = disable, 0 = enable)
            CM06 : Bool;   // CMxx (1 = disable, 0 = enable)
            CM07 : Bool;   // CMxx (1 = disable, 0 = enable)
            CM08 : Bool;   // CMxx (1 = disable, 0 = enable)
            CM09 : Bool;   // CMxx (1 = disable, 0 = enable)
            CM10 : Bool;   // CMxx (1 = disable, 0 = enable)
         END_STRUCT;
      END_STRUCT;
   END_VAR
BEGIN
   Names.statesNames[1,1] := 'Clearing';
   Names.statesNames[1,2] := 'Stopped';
   Names.statesNames[1,3] := 'Starting';
   Names.statesNames[1,4] := 'Idle';
   Names.statesNames[1,5] := 'Suspended';
   Names.statesNames[1,6] := 'Execute';
   Names.statesNames[1,7] := 'Stopping';
   Names.statesNames[1,8] := 'Aborting';
   Names.statesNames[1,9] := 'Aborted';
   Names.statesNames[1,10] := 'Holding';
   Names.statesNames[1,11] := 'Held';
   Names.statesNames[1,12] := 'UnHolding';
   Names.statesNames[1,13] := 'Suspending';
   Names.statesNames[1,14] := 'UnSuspending';
   Names.statesNames[1,15] := 'Resetting';
   Names.statesNames[1,16] := 'Completing';
   Names.statesNames[1,17] := 'Complete';
   Names.unitModesNames[2,0] := 'Invalid';
   Names.unitModesNames[2,1] := 'Production';
   Names.unitModesNames[2,2] := 'Maintenance';
   Names.unitModesNames[2,3] := 'Manual';
   Names.unitModesNames[2,4] := 'User Mode 01';
   Names.statesNames[2,1] := 'Limpiar';
   Names.statesNames[2,2] := 'Detenido';
   Names.statesNames[2,3] := 'Empezando';
   Names.statesNames[2,4] := 'Parado';
   Names.statesNames[2,5] := 'Interrumpido';
   Names.statesNames[2,6] := 'Correr';
   Names.statesNames[2,7] := 'Detener';
   Names.statesNames[2,8] := 'Anulando';
   Names.statesNames[2,9] := 'Anulado';
   Names.statesNames[2,10] := 'Mantener';
   Names.statesNames[2,11] := 'Mantenido';
   Names.statesNames[2,12] := 'Desmentener';
   Names.statesNames[2,13] := 'Interrumpir';
   Names.statesNames[2,14] := 'Desinterrumpir';
   Names.statesNames[2,15] := 'Reajustar';
   Names.statesNames[2,16] := 'Terminar';
   Names.statesNames[2,17] := 'Terminado';
   Names.statesNames[2,0] := 'Undefined';
END_DATA_BLOCK

